// TIA Portal project "test_program" (V15)

(* hardware
DEVICE "S71500/ET200MP station_1"  S7-1500 station
   slot 0: "Rail_0"  Rack  6ES7 590-1***0-0AA0
   slot 0: "PS 25W 24VDC_1"  PS 25W 24VDC  6ES7 505-0KA00-0AB0  V1.0
   slot 1: "PLC_1"  CPU 1511F-1 PN  6ES7 511-1FK01-0AB0  V1.8
   slot 2: "DI 16x24VDC HF_1"  DI 16x24VDC HF  6ES7 521-1BH00-0AB0  V2.0
   slot 3: "DI 16x24VDC HF_2"  DI 16x24VDC HF  6ES7 521-1BH00-0AB0  V2.0
   slot 4: "AI 8xU/I/RTD/TC ST_1"  AI 8xU/I/RTD/TC ST  6ES7 531-7KF00-0AB0  V2.1
DEVICE "SCALANCE X005"  SCALANCE X-Station
   slot 0: "SCALANCE X rack"  Rail
   slot 0: "Switch_1"  6GK5 005-0BA00-1AA3  V1.0
*)

// ===== PLC "PLC_1"  CPU 1511F-1 PN =====
// protected blocks, not shown: "Main_Safety_RTG1_1", "Main_Safety_RTG1_DB_1"

TYPE "Drive_To_PLC"
   STRUCT
      IN_DI1_Enable_status : Bool;
      IN_DI2_Drive_error : Bool;
      IN_DI3 : Bool;
      IN_DI4 : Bool;
      IN_AI1_Pressure_feedback : UInt;
      IN_AI2_Flow_feedback : UInt;
   END_STRUCT;
END_TYPE

TYPE "PLC_To_Drive"
   STRUCT
      OUT_DO1_Enable : Bool;
      OUT_DO2_PID_gain_select : Bool;
      OUT_DO3_Slave_select : Bool;
      OUT_DO4_Fault_reset : Bool;
      OUT_DO5_CAN_comm_enable : Bool;
      OUT_AO1_Pressure_command : UInt;
      OUT_AO2_Flow_command : UInt;
   END_STRUCT;
END_TYPE

DATA_BLOCK "Inputs_DB"   // DB2
{ S7_Optimized_Access := 'TRUE' }
VERSION : 0.1
   VAR
      Immediate_STOP : Bool;
      Reset : Bool;
   END_VAR
BEGIN
END_DATA_BLOCK

DATA_BLOCK "Outputs_DB"   // DB3
{ S7_Optimized_Access := 'TRUE' }
VERSION : 0.1
BEGIN
END_DATA_BLOCK

// folder: IS580_HydraulicServoDrive

DATA_BLOCK "IS580_HydraulicServoDrive_Control_DB"   // DB100
{ S7_Optimized_Access := 'TRUE' }
VERSION : 0.1
   VAR
      Pressure_SETPOINT : Real;
      FLow_SETPOINT : Real;
      Pressure_FEEDBACK : Real;
      FLow_FEEDBACK : Real;
      PI : "Drive_To_PLC";
      PO : "PLC_To_Drive";
   END_VAR
BEGIN
END_DATA_BLOCK

// folder: (top level)

FUNCTION "SCALE_UInt_TO_REAL" : Void   // FC700, FBD
TITLE = Scaling_Function_2
{ S7_Optimized_Access := 'TRUE' }
VERSION : 0.1
   VAR_INPUT
      Input_Min : Real;
      Input_Max : Int;
      Input_Signal : Real;
      Output_Min : Real;
      Output_Max : Real;
   END_VAR
   VAR_OUTPUT
      SV : Real;
   END_VAR
   VAR_TEMP
      tv : Real;
   END_VAR
BEGIN

REGION Network 1
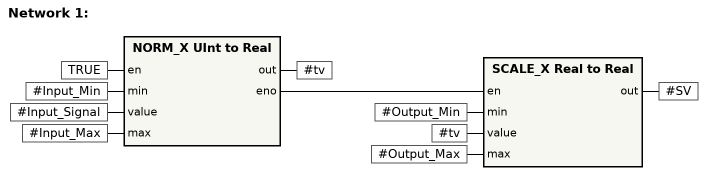
   IF TRUE THEN
       #tv := NORM_X(MIN := #Input_Min, VALUE := #Input_Signal, MAX := #Input_Max);
       #SV := SCALE_X(MIN := #Output_Min, VALUE := #tv, MAX := #Output_Max);
   END_IF;
END_REGION
END_FUNCTION

FUNCTION "SCALE_REAL_TO_UInt" : Void   // FC701, FBD
TITLE = Scaling_Function_2
{ S7_Optimized_Access := 'TRUE' }
VERSION : 0.1
   VAR_INPUT
      Input_Min : Real;
      Input_Max : Int;
      Input_Signal : Real;
      Output_Min : Real;
      Output_Max : Real;
   END_VAR
   VAR_OUTPUT
      SV : UInt;
   END_VAR
   VAR_TEMP
      tv : Real;
   END_VAR
BEGIN

REGION Network 1
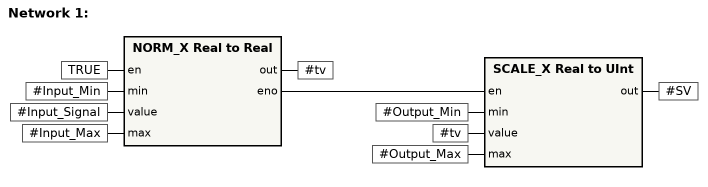
   IF TRUE THEN
       #tv := NORM_X(MIN := #Input_Min, VALUE := #Input_Signal, MAX := #Input_Max);
       #SV := SCALE_X(MIN := #Output_Min, VALUE := #tv, MAX := #Output_Max);
   END_IF;
END_REGION
END_FUNCTION

ORGANIZATION_BLOCK "Main"   // OB1, LAD, ProgramCycle
TITLE = "Main Program Sweep (Cycle)"
{ S7_Optimized_Access := 'TRUE' }
VERSION : 0.1
   VAR_INPUT
      Initial_Call : Bool;   // Initial call of this OB
      Remanence : Bool;   // =True, if remanent data are available
   END_VAR
   VAR_TEMP
      "Abort_with_SS (Auto to Manual)" : Bool;
      "Abort_with_SS (Manual to Auto)" : Bool;
      Initialize_Graph_Manual_Cycle : Bool;
      Abort_Cycle_Common_bit : Bool;
      TX_Recipe_Transfer : Bool;
      Blk_Return_P1 : Int;
      Blk_Return_P2 : Int;
      Blk_Return_P3 : Int;
      Blk_Return_P4 : Int;
      Blk_Return_P5 : Int;
      Blk_Return_P6 : Int;
      Blk_Return_P7 : Int;
      Blk_Return_P8 : Int;
      Blk_Return_P9 : Int;
   END_VAR
BEGIN

REGION Network 1
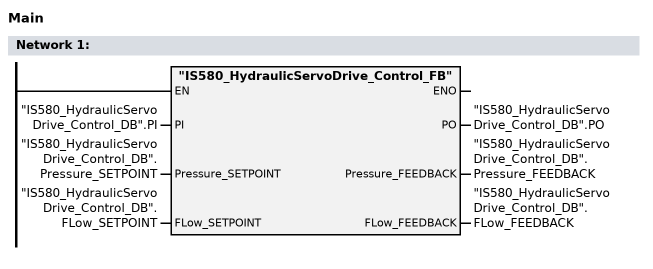
   RUNG wire#powerrail
      "IS580_HydraulicServoDrive_Control_FB"(PI := "IS580_HydraulicServoDrive_Control_DB".PI, PO => "IS580_HydraulicServoDrive_Control_DB".PO, Pressure_SETPOINT := "IS580_HydraulicServoDrive_Control_DB".Pressure_SETPOINT, FLow_SETPOINT := "IS580_HydraulicServoDrive_Control_DB".FLow_SETPOINT, Pressure_FEEDBACK => "IS580_HydraulicServoDrive_Control_DB".Pressure_FEEDBACK, FLow_FEEDBACK => "IS580_HydraulicServoDrive_Control_DB".FLow_FEEDBACK)
   END_RUNG
   // the same network as SCL:
   "IS580_HydraulicServoDrive_Control_FB"(PI := "IS580_HydraulicServoDrive_Control_DB".PI,
                           Pressure_SETPOINT := "IS580_HydraulicServoDrive_Control_DB".Pressure_SETPOINT,
                           FLow_SETPOINT := "IS580_HydraulicServoDrive_Control_DB".FLow_SETPOINT,
                           PO => "IS580_HydraulicServoDrive_Control_DB".PO,
                           Pressure_FEEDBACK => "IS580_HydraulicServoDrive_Control_DB".Pressure_FEEDBACK,
                           FLow_FEEDBACK => "IS580_HydraulicServoDrive_Control_DB".FLow_FEEDBACK);
END_REGION
END_ORGANIZATION_BLOCK

// folder: IS580_HydraulicServoDrive

FUNCTION "IS580_HydraulicServoDrive_Control_FB" : Void   // FC100, SCL
{ S7_Optimized_Access := 'TRUE' }
VERSION : 0.1
   VAR_INPUT
      PI : "Drive_To_PLC";
      Pressure_SETPOINT : Real;
      FLow_SETPOINT : Real;
   END_VAR
   VAR_OUTPUT
      PO : "PLC_To_Drive";
      Pressure_FEEDBACK : Real;
      FLow_FEEDBACK : Real;
   END_VAR
BEGIN
   (*
   Suppose we have a hydraulic system where the MAX/MIN limit are as following
   MAX_Pressure = 320 bar
   MIN_Pressure = 0 bar
   MAX_Flow = 20 L/min
   MIN_Flow = 0 L/min
   Pressure & Flow command to the Inverter are given within these limits
   *)

   //***************************************************
   IF  "Inputs_DB".Immediate_STOP = FALSE
       AND #PI.IN_DI2_Drive_error = FALSE
       AND "IS580_HydraulicServoDrive_Control_DB".PI.IN_DI1_Enable_status = TRUE THEN
       //Pressure command
       "SCALE_REAL_TO_UInt"(Input_Min := 0,
                            Input_Max := 320,
                            Input_Signal := #Pressure_SETPOINT,
                            Output_Min := 0.0,
                            Output_Max := 27648,
                            SV => #PO.OUT_AO1_Pressure_command);
       //Flow command
       "SCALE_REAL_TO_UInt"(Input_Min:=0,
                            Input_Max:=20,
                            Input_Signal:=#FLow_SETPOINT,
                            Output_Min:=0,
                            Output_Max:=27648,
                            SV=>#PO.OUT_AO2_Flow_command);

   ELSE
       //Pressure command > Null
       "SCALE_REAL_TO_UInt"(Input_Min := 0,
                            Input_Max := 100,
                            Input_Signal := 0.0,
                            Output_Min := 0.0,
                            Output_Max := 27648,
                            SV => #PO.OUT_AO1_Pressure_command);
       //Flow command > Null
       "SCALE_REAL_TO_UInt"(Input_Min := 0,
                            Input_Max := 250,
                            Input_Signal := 0.0,
                            Output_Min := 0,
                            Output_Max := 27648,
                            SV => #PO.OUT_AO2_Flow_command);
   END_IF;

   //***************************************************
   //Pressure feedback
   "SCALE_UInt_TO_REAL"(Input_Min:=0,
                        Input_Max:=27648,
                        Input_Signal:=#PI.IN_AI1_Pressure_feedback,
                        Output_Min:=0.0,
                        Output_Max:=100.0,
                        SV=>#Pressure_FEEDBACK);

   //Flow feedback
   "SCALE_UInt_TO_REAL"(Input_Min:=0,
                        Input_Max:=27648,
                        Input_Signal:=#PI.IN_AI2_Flow_feedback,
                        Output_Min:=0.0,
                        Output_Max:=250.0,
                        SV=>#FLow_FEEDBACK);

   //***************************************************
   //Inverter fault reset
   #PO.OUT_DO4_Fault_reset := "Inputs_DB".Reset;
END_FUNCTION